VERSION : 0.1
   VAR_INPUT
      CMD : Bool;   // Команда запуска
      Res_1 : DInt;   // Наработка устройства 1
      Res_2 : DInt;   // Наработка устройства 2
      Alm_1 : Bool;   // Авария устройства 1
      Alm_2 : Bool;   // Авария устройства 2
   END_VAR
   VAR_IN_OUT
      Res_SP : DInt;   // Переключение по наработке
      CMD_1 : Bool;   // Команда на устройство 1
      CMD_2 : Bool;   // Команда на устройство 2
   END_VAR
   VAR_TEMP
      N : Bool;   // Выбор устройства
      Now : DInt;   // Текущая разница наработок
   END_VAR
BEGIN

REGION Network 1: Подсчёт разницы наработки
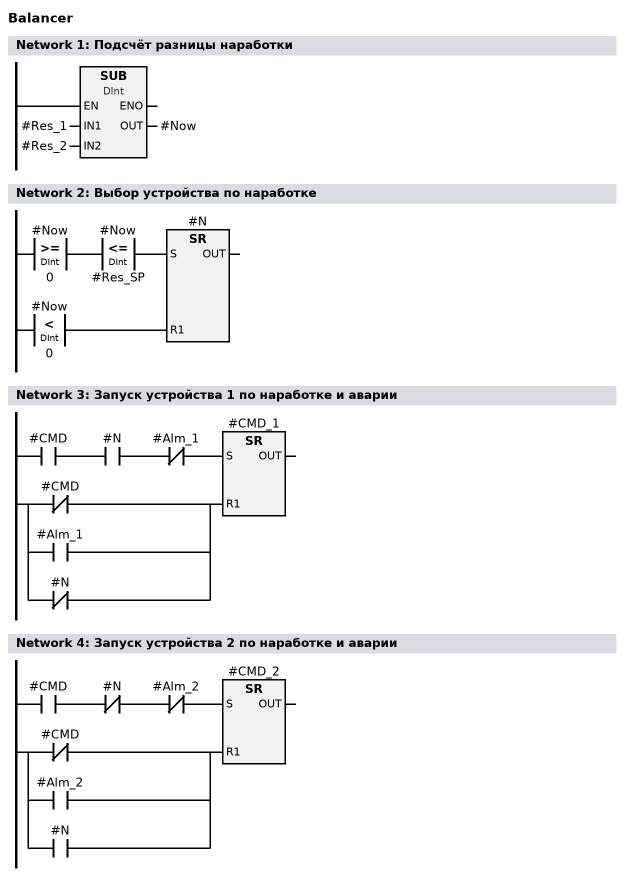
   RUNG wire#powerrail
      { S7_Templates := "SrcType := DInt"; S7_GenerateENO := "TRUE" } Sub(in1 := #Res_1, in2 := #Res_2, out => #Now)
   END_RUNG
   // the same network as SCL:
   #Now := #Res_1 - #Res_2;
END_REGION

REGION Network 2: Выбор устройства по наработке
   RUNG wire#powerrail
      { S7_Templates := "SrcType := DInt" } GE_Contact(in1 := #Now, in2 := 0)
      { S7_Templates := "SrcType := DInt" } LE_Contact(in1 := #Now, in2 := #Res_SP)
      S_SR(operand := #N, r1 := wire#w1)
   END_RUNG
   RUNG wire#powerrail
      { S7_Templates := "SrcType := DInt" } LT_Contact(in1 := #Now, in2 := 0)
   END_RUNG wire#w1
   // the same network as SCL:
   IF (#Now >= 0) AND (#Now <= #Res_SP) THEN
       #N := TRUE;   // SR flip-flop
   END_IF;
   IF #Now < 0 THEN #N := FALSE; END_IF;
END_REGION

REGION Network 3: Запуск устройства 1 по наработке и аварии
   RUNG wire#powerrail
      Contact( #CMD )
      Contact( #N )
      I_Contact( #Alm_1 )
      S_SR(operand := #CMD_1, r1 := wire#w1)
   END_RUNG
   RUNG wire#powerrail
      I_Contact( #CMD )
   END_RUNG wire#w1
   RUNG wire#powerrail
      Contact( #Alm_1 )
   END_RUNG wire#w1
   RUNG wire#powerrail
      I_Contact( #N )
   END_RUNG wire#w1
   // the same network as SCL:
   IF #CMD AND #N AND NOT #Alm_1 THEN
       #CMD_1 := TRUE;   // SR flip-flop
   END_IF;
   IF NOT #CMD OR #Alm_1 OR NOT #N THEN #CMD_1 := FALSE; END_IF;
END_REGION

REGION Network 4: Запуск устройства 2 по наработке и аварии
   RUNG wire#powerrail
      Contact( #CMD )
      I_Contact( #N )
      I_Contact( #Alm_2 )
      S_SR(operand := #CMD_2, r1 := wire#w1)
   END_RUNG
   RUNG wire#powerrail
      I_Contact( #CMD )
   END_RUNG wire#w1
   RUNG wire#powerrail
      Contact( #Alm_2 )
   END_RUNG wire#w1
   RUNG wire#powerrail
      Contact( #N )
   END_RUNG wire#w1
   // the same network as SCL:
   IF #CMD AND NOT #N AND NOT #Alm_2 THEN
       #CMD_2 := TRUE;   // SR flip-flop
   END_IF;
   IF NOT #CMD OR #Alm_2 OR #N THEN #CMD_2 := FALSE; END_IF;
END_REGION
END_FUNCTION

FUNCTION "INV" : Void   // FC111, LAD
{ S7_Optimized_Access := 'TRUE' }
VERSION : 0.1
   VAR_INPUT
      S : Bool;   // Сигнал
      I : Bool;   // Инверсия
   END_VAR
   VAR_IN_OUT
      R : Bool;   // Результат
   END_VAR
BEGIN

REGION Network 1: Инверсия сигнала
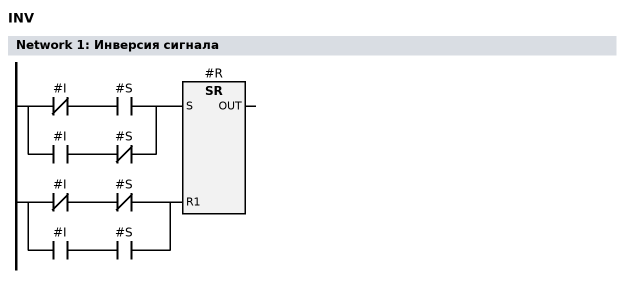
   RUNG wire#powerrail
      I_Contact( #I )
      Contact( #S )
      wire#w1
      S_SR(operand := #R, r1 := wire#w2)
   END_RUNG
   RUNG wire#powerrail
      Contact( #I )
      I_Contact( #S )
   END_RUNG wire#w1
   RUNG wire#powerrail
      I_Contact( #I )
      I_Contact( #S )
   END_RUNG wire#w2
   RUNG wire#powerrail
      Contact( #I )
      Contact( #S )
   END_RUNG wire#w2
   // the same network as SCL:
   IF (NOT #I AND #S) OR (#I AND NOT #S) THEN
       #R := TRUE;   // SR flip-flop
   END_IF;
   IF (NOT #I AND NOT #S) OR (#I AND #S) THEN #R := FALSE; END_IF;
END_REGION
END_FUNCTION

FUNCTION "Mode" : Void   // FC150, LAD
{ S7_Optimized_Access := 'FALSE' }
VERSION : 0.1
   VAR_INPUT
      CMD : Struct   // Основные команды
         Hand : Bool;   // 0 - авто, 1 - ручной / 0 - Авто, 1 - Ручной
         Start_A : Bool;   // Автозапуск / Запуск в авторежиме
         Start_M : Bool;   // Ручной - вперёд / Запуск в ручном режиме
         Force : Bool;   // Принудительный
         Lock : Bool;   // Блокировать / Блокировка
         Local : Bool;   // Локальный
         Service : Bool;   // Сервис
         Safety : Bool;   // Безопасность
         Alarm : Bool;   // Есть авария / Авария
         Reset : Bool;   // Сброс аварий
         Sim : Bool;   // Режим симуляции
      END_STRUCT;
      All_Block : Bool;   // Аварийная блокировка
   END_VAR
   VAR_OUTPUT
      Mode : Int;   // Режим работы
   END_VAR
BEGIN

REGION Network 1: Автоматический режим
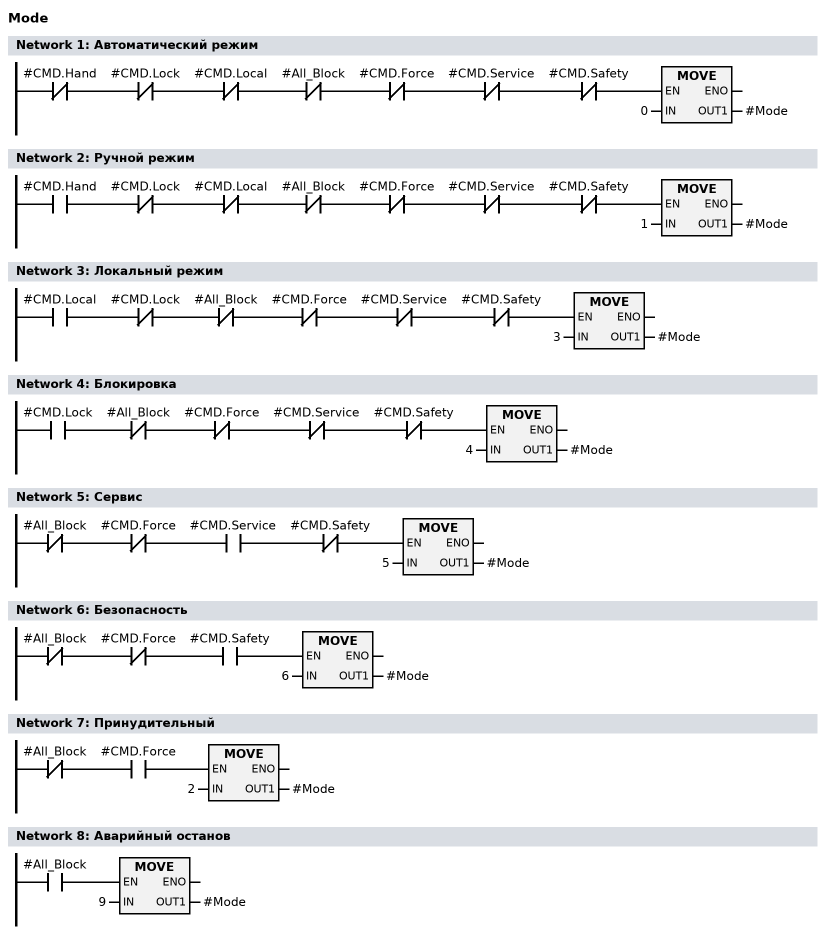
   RUNG wire#powerrail
      I_Contact( #CMD.Hand )
      I_Contact( #CMD.Lock )
      I_Contact( #CMD.Local )
      I_Contact( #All_Block )
      I_Contact( #CMD.Force )
      I_Contact( #CMD.Service )
      I_Contact( #CMD.Safety )
      { S7_GenerateENO := "TRUE" } Move(in := 0, out1 => #Mode)
   END_RUNG
   // the same network as SCL:
   IF NOT #CMD.Hand AND NOT #CMD.Lock AND NOT #CMD.Local AND NOT #All_Block AND NOT #CMD.Force AND NOT #CMD.Service AND NOT #CMD.Safety THEN
       #Mode := 0;
   END_IF;
END_REGION

REGION Network 2: Ручной режим
   RUNG wire#powerrail
      Contact( #CMD.Hand )
      I_Contact( #CMD.Lock )
      I_Contact( #CMD.Local )
      I_Contact( #All_Block )
      I_Contact( #CMD.Force )
      I_Contact( #CMD.Service )
      I_Contact( #CMD.Safety )
      { S7_GenerateENO := "TRUE" } Move(in := 1, out1 => #Mode)
   END_RUNG
   // the same network as SCL:
   IF #CMD.Hand AND NOT #CMD.Lock AND NOT #CMD.Local AND NOT #All_Block AND NOT #CMD.Force AND NOT #CMD.Service AND NOT #CMD.Safety THEN
       #Mode := 1;
   END_IF;
END_REGION

REGION Network 3: Локальный режим
   RUNG wire#powerrail
      Contact( #CMD.Local )
      I_Contact( #CMD.Lock )
      I_Contact( #All_Block )
      I_Contact( #CMD.Force )
      I_Contact( #CMD.Service )
      I_Contact( #CMD.Safety )
      { S7_GenerateENO := "TRUE" } Move(in := 3, out1 => #Mode)
   END_RUNG
   // the same network as SCL:
   IF #CMD.Local AND NOT #CMD.Lock AND NOT #All_Block AND NOT #CMD.Force AND NOT #CMD.Service AND NOT #CMD.Safety THEN
       #Mode := 3;
   END_IF;
END_REGION

REGION Network 4: Блокировка
   RUNG wire#powerrail
      Contact( #CMD.Lock )
      I_Contact( #All_Block )
      I_Contact( #CMD.Force )
      I_Contact( #CMD.Service )
      I_Contact( #CMD.Safety )
      { S7_GenerateENO := "TRUE" } Move(in := 4, out1 => #Mode)
   END_RUNG
   // the same network as SCL:
   IF #CMD.Lock AND NOT #All_Block AND NOT #CMD.Force AND NOT #CMD.Service AND NOT #CMD.Safety THEN
       #Mode := 4;
   END_IF;
END_REGION

REGION Network 5: Сервис
   RUNG wire#powerrail
      I_Contact( #All_Block )
      I_Contact( #CMD.Force )
      Contact( #CMD.Service )
      I_Contact( #CMD.Safety )
      { S7_GenerateENO := "TRUE" } Move(in := 5, out1 => #Mode)
   END_RUNG
   // the same network as SCL:
   IF NOT #All_Block AND NOT #CMD.Force AND #CMD.Service AND NOT #CMD.Safety THEN #Mode := 5; END_IF;
END_REGION

REGION Network 6: Безопасность
   RUNG wire#powerrail
      I_Contact( #All_Block )
      I_Contact( #CMD.Force )
      Contact( #CMD.Safety )
      { S7_GenerateENO := "TRUE" } Move(in := 6, out1 => #Mode)
   END_RUNG
   // the same network as SCL:
   IF NOT #All_Block AND NOT #CMD.Force AND #CMD.Safety THEN #Mode := 6; END_IF;
END_REGION

REGION Network 7: Принудительный
   RUNG wire#powerrail
      I_Contact( #All_Block )
      Contact( #CMD.Force )
      { S7_GenerateENO := "TRUE" } Move(in := 2, out1 => #Mode)
   END_RUNG
   // the same network as SCL:
   IF NOT #All_Block AND #CMD.Force THEN #Mode := 2; END_IF;
END_REGION

REGION Network 8: Аварийный останов
   RUNG wire#powerrail
      Contact( #All_Block )
      { S7_GenerateENO := "TRUE" } Move(in := 9, out1 => #Mode)
   END_RUNG
   // the same network as SCL:
   IF #All_Block THEN #Mode := 9; END_IF;
END_REGION
END_FUNCTION

// ===== PLC "PLC_PolyMix_002"  CPU 1214C DC/DC/DC =====
// protected blocks, not shown: "AI_ex", "AIx", "AO_ex", "DRV_M_D", "FlowMeter", "Logick", "Motors", "PLF_FC", "Time_m", "Time_r", "Time_s"

VAR_GLOBAL   // PLC tag table "Default tag table"
   "Mix_1_Clock" AT %M10.0 : Bool;
   "Mix_2_Clock" AT %M10.1 : Bool;
   "Mix_3_Clock" AT %M10.2 : Bool;
   "Flow" AT %IW256 : Int;
   "Level" AT %IW258 : Int;
END_VAR

VAR_GLOBAL   // PLC tag table "Sys"
   "pulse_01s" AT %M2.0 : Bool;
   "pulse_05s" AT %M2.1 : Bool;
   "pulse_1s" AT %M2.2 : Bool;
   "All_block" AT %M3.0 : Bool;
   "Reset_All" AT %M3.1 : Bool;
   "Sim_All" AT %M3.2 : Bool;
   "Any_Hand" AT %M5.0 : Bool;
   "DI_Hand" AT %M5.1 : Bool;
   "DO_Hand" AT %M5.2 : Bool;
   "AI_Hand" AT %M5.3 : Bool;
   "AO_Hand" AT %M5.4 : Bool;
   "M_Hand" AT %M5.5 : Bool;
   "V_Hand" AT %M5.6 : Bool;
   "X_Hand" AT %M5.7 : Bool;
   "System_Byte" AT %MB1 : Byte;
   "FirstScan" AT %M1.0 : Bool;
   "DiagStatusUpdate" AT %M1.1 : Bool;
   "ON" AT %M1.2 : Bool;
   "OFF" AT %M1.3 : Bool;
   "Clock_Byte" AT %MB0 : Byte;
   "Clock_10Hz" AT %M0.0 : Bool;
   "Clock_5Hz" AT %M0.1 : Bool;
   "Clock_2.5Hz" AT %M0.2 : Bool;
   "Clock_2Hz" AT %M0.3 : Bool;
   "Clock_1.25Hz" AT %M0.4 : Bool;
   "Clock_1Hz" AT %M0.5 : Bool;
   "Clock_0.625Hz" AT %M0.6 : Bool;
   "Clock_0.5Hz" AT %M0.7 : Bool;
   "F_pulse_01s" AT %M2.3 : Bool;
   "F_pulse_05s" AT %M2.4 : Bool;
   "F_pulse_1s" AT %M2.5 : Bool;
   "FN_pulse_01s" AT %M2.6 : Bool;
   "Clock_5s" AT %M2.7 : Bool;
   "Any_Alm" AT %M6.0 : Bool;
   "AI_Alm" AT %M6.1 : Bool;
   "M_Alm" AT %M6.2 : Bool;
   "V_Alm" AT %M6.3 : Bool;
   "C_Alm" AT %M6.4 : Bool;
   "N_Alm" AT %M6.5 : Bool;
   "L_Alm" AT %M6.6 : Bool;
   "X_Alm" AT %M6.7 : Bool;
END_VAR

VAR_GLOBAL   // PLC tag table "IO Table"
   "DD_FB_Ready" AT %I0.6 : Bool;   // I 0.6 - Дозатор сухого вещества - готовность
   "Dos_FB_Run" AT %I0.7 : Bool;   // I 0.7 - Дозатор - работа
   "DD_LLS" AT %I1.0 : Bool;   // I 1.0 - Дозатор сухого вещества - низкий уровень
   "Vibro_FB_Ready" AT %I1.1 : Bool;   // I 1.1 - Вибратор - готовность
   "Transporter" AT %I1.2 : Bool;   // I 1.2 - Пневмотранспортёр - готовность
   "DL_FB_Ready" AT %I1.3 : Bool;   // I 1.3 - Дозатор жидкого вещества - готовность
   "Dry_Run" AT %I1.4 : Bool;   // I 1.4 - Датчик протока
   "AllBlock" AT %I1.5 : Bool;   // I 1.5 - Датчик перелива или Аварийная остановка
   "M1_FB_Ready" AT %I0.0 : Bool;   // I 0.0 - Мешалка 1 - готовность
   "M1_FB_Run" AT %I0.1 : Bool;   // I 0.1 - Мешалка 1 - работа
   "M2_FB_Ready" AT %I0.2 : Bool;   // I 0.2 - Мешалка 2 - готовность
   "M2_FB_Run" AT %I0.3 : Bool;   // I 0.3 - Мешалка 2 - работа
   "M3_FB_Ready" AT %I0.4 : Bool;   // I 0.4 - Мешалка 3 - готовность
   "M3_FB_Run" AT %I0.5 : Bool;   // I 0.5 - Мешалка 3 - работа
   "M1_CMD" AT %Q0.0 : Bool;   // Q 0.0 - Мешалка 1 - запуск
   "M2_CMD" AT %Q0.1 : Bool;   // Q 0.1 - Мешалка 2 - запуск
   "M3_CMD" AT %Q0.2 : Bool;   // Q 0.2 - Мешалка 3 - запуск
   "DD_CMD" AT %Q0.3 : Bool;   // Q 0.3 - Дозатор сухого вещества - запуск
   "Vibro_CMD" AT %Q0.4 : Bool;   // Q 0.4 - Вибратор - запуск
   "DL_CMD" AT %Q0.5 : Bool;   // Q 0.5 - Дозатор жидкого вещества - запуск
   "KC1_CMD" AT %Q0.6 : Bool;   // Q 0.6 - Соленоидный клапан КС1
   "LED_Dry_Run" AT %Q0.7 : Bool;   // Q 0.7 - LED - сухой ход
   "LED_Alarm" AT %Q1.0 : Bool;   // Q 1.0 - LED - общая авария
   "LED_Empty" AT %Q1.1 : Bool;   // Q 1.1 - LED - бункер пуст
END_VAR

DATA_BLOCK "Any_DB"   // DB3
{ S7_Optimized_Access := 'FALSE' }
VERSION : 0.1
   VAR
      Level_M : Int;
      Level_S : Int;
      Flow_M : Int;
      Flow_S : Int;
      DD_View : Bool;
      Level_View : Bool;
   END_VAR
BEGIN
END_DATA_BLOCK

DATA_BLOCK "CONFIG"   // DB10
{ S7_Optimized_Access := 'FALSE' }
VERSION : 0.1
   VAR
      Config : Struct
         Use_DD : Bool;   // Использовать сухой дозатор
         Use_DL : Bool := true;   // Использовать жидкий дозатор
         Use_Mix_1 : Bool := true;   // Использовать мешалку 1
         Use_Mix_2 : Bool := true;   // Использовать мешалку 2
         Use_Mix_3 : Bool := true;   // Использовать мешалку 3
      END_STRUCT;
   END_VAR
BEGIN
END_DATA_BLOCK

DATA_BLOCK "Comm_DB"   // DB11
{ S7_Optimized_Access := 'FALSE' }
VERSION : 0.1
   VAR
      DD_Status : Int;
      DD_Mode : Int;
      DD_Alarm : Word;
      DL_Status : Int;
      DL_Mode : Int;
      DL_Alarm : Word;
      Mix_1_Status : Int;
      Mix_1_Mode : Int;
      Mix_1_Alarm : Word;
      Mix_2_Status : Int;
      Mix_2_Mode : Int;
      Mix_2_Alarm : Word;
      Mix_3_Status : Int;
      Mix_3_Mode : Int;
      Mix_3_Alarm : Word;
      KC1_Status : Int;
      Flowmeter : Real;
      Flow_Alarm : Word;
      Level : Real;
      Level_Alarm : Word;
      SP : Real;
      Start : Bool;
      Hand : Bool;
      Warning : Bool;
      Config : Struct
         Use_DD : Bool;   // Использовать сухой дозатор
         Use_DL : Bool;   // Использовать жидкий дозатор
         Use_Mix_1 : Bool;   // Использовать мешалку 1
         Use_Mix_2 : Bool;   // Использовать мешалку 2
         Use_Mix_3 : Bool;   // Использовать мешалку 3
      END_STRUCT;
      Alarm : Word;
   END_VAR
BEGIN
END_DATA_BLOCK

// folder: Modules

DATA_BLOCK "DIx_DB"   // DB200
{ S7_Optimized_Access := 'FALSE' }
VERSION : 0.1
// stored: InstanceOfName DIx
"DIx"
BEGIN
END_DATA_BLOCK

DATA_BLOCK "DOx_DB"   // DB201
{ S7_Optimized_Access := 'FALSE' }
VERSION : 0.1
// stored: InstanceOfName DOx
"DOx"
BEGIN
END_DATA_BLOCK

DATA_BLOCK "Micro_DB"   // DB207
{ S7_Optimized_Access := 'FALSE' }
VERSION : 0.1
// stored: InstanceOfName Micro
"Micro"
BEGIN
END_DATA_BLOCK

// folder: System blocks/Program resources

DATA_BLOCK "T_Reset"   // DB7
{ S7_Optimized_Access := 'TRUE' }
AUTHOR : Simatic
FAMILY : IEC
NAME : IEC_TMR
VERSION : 1.0
// stored: InstanceOfName IEC_TIMER
"IEC_TIMER"
BEGIN
END_DATA_BLOCK

DATA_BLOCK "clock_5s_ON"   // DB507
{ S7_Optimized_Access := 'TRUE' }
AUTHOR : Simatic
FAMILY : IEC
NAME : IEC_TMR
VERSION : 1.0
// stored: InstanceOfName IEC_TIMER
"IEC_TIMER"
BEGIN
END_DATA_BLOCK

DATA_BLOCK "clock_5s_OFF"   // DB508
{ S7_Optimized_Access := 'TRUE' }
AUTHOR : Simatic
FAMILY : IEC
NAME : IEC_TMR
VERSION : 1.0
// stored: InstanceOfName IEC_TIMER
"IEC_TIMER"
BEGIN
END_DATA_BLOCK

// folder: (top level)

FUNCTION "Comm_FC" : Void   // FC1, LAD
{ S7_Optimized_Access := 'TRUE' }
VERSION : 0.1
BEGIN

REGION Network 1: Сухой дозатор
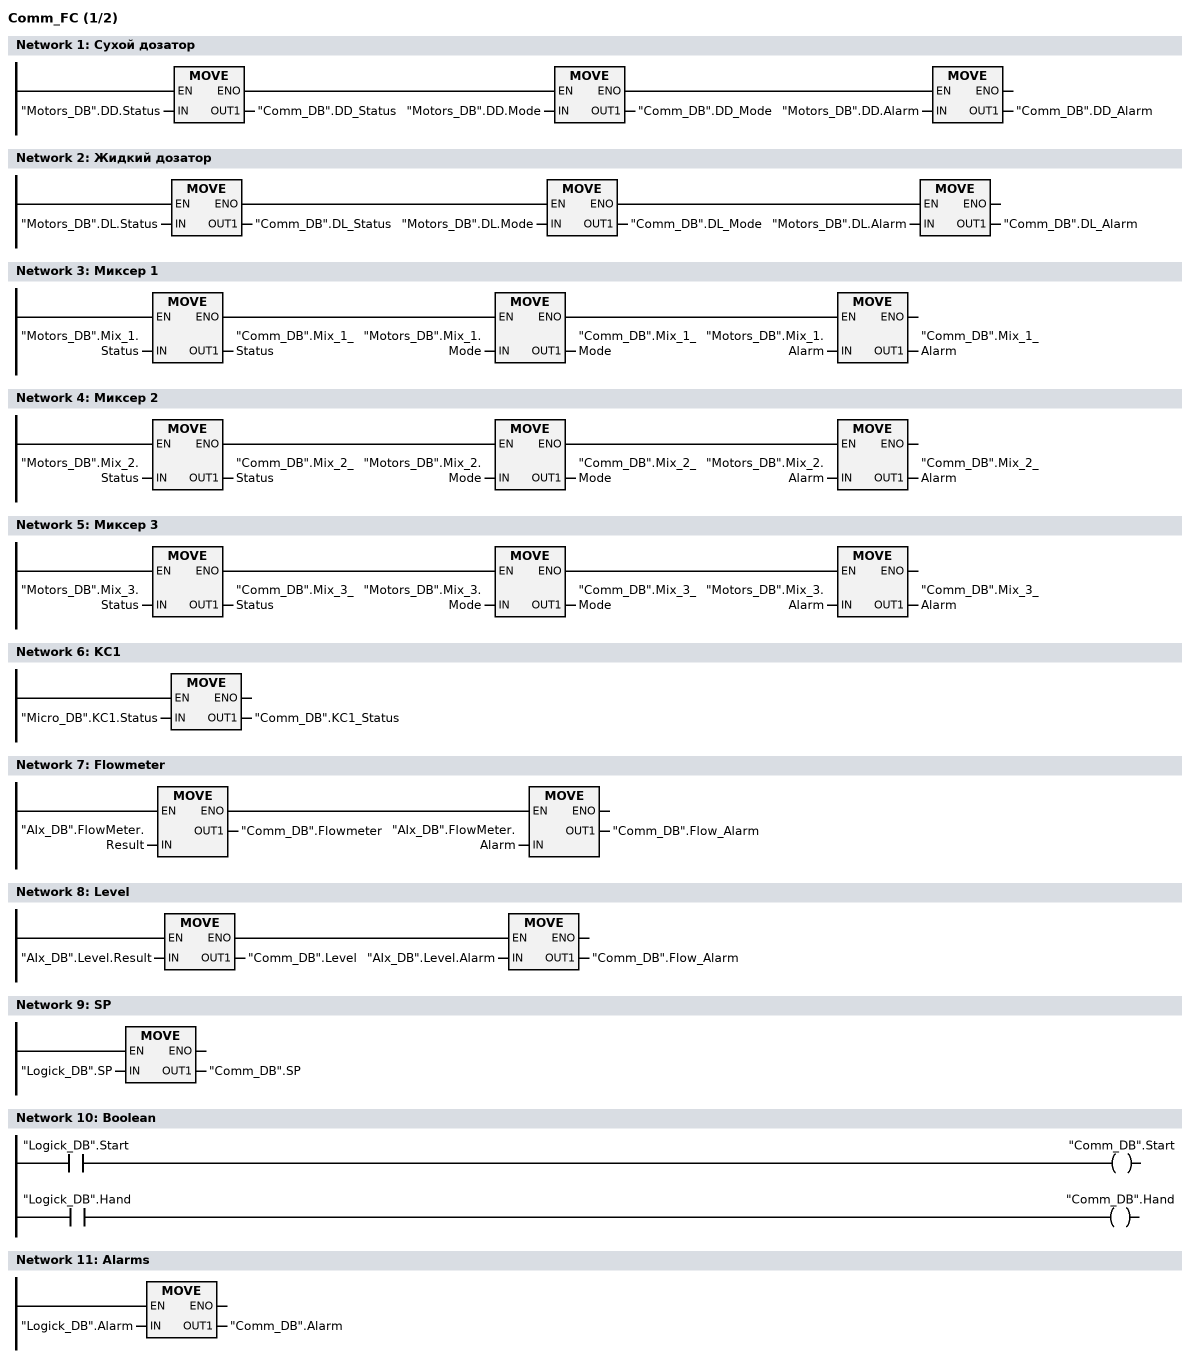
   RUNG wire#powerrail
      Move(in := "Motors_DB".DD.Status, out1 => "Comm_DB".DD_Status)
      Move(in := "Motors_DB".DD.Mode, out1 => "Comm_DB".DD_Mode)
      Move(in := "Motors_DB".DD.Alarm, out1 => "Comm_DB".DD_Alarm)
   END_RUNG
   // the same network as SCL:
   "Comm_DB".DD_Status := "Motors_DB".DD.Status;
   "Comm_DB".DD_Mode := "Motors_DB".DD.Mode;
   "Comm_DB".DD_Alarm := "Motors_DB".DD.Alarm;
END_REGION

REGION Network 2: Жидкий дозатор
   RUNG wire#powerrail
      Move(in := "Motors_DB".DL.Status, out1 => "Comm_DB".DL_Status)
      Move(in := "Motors_DB".DL.Mode, out1 => "Comm_DB".DL_Mode)
      Move(in := "Motors_DB".DL.Alarm, out1 => "Comm_DB".DL_Alarm)
   END_RUNG
   // the same network as SCL:
   "Comm_DB".DL_Status := "Motors_DB".DL.Status;
   "Comm_DB".DL_Mode := "Motors_DB".DL.Mode;
   "Comm_DB".DL_Alarm := "Motors_DB".DL.Alarm;
END_REGION

REGION Network 3: Миксер 1
   RUNG wire#powerrail
      Move(in := "Motors_DB".Mix_1.Status, out1 => "Comm_DB".Mix_1_Status)
      Move(in := "Motors_DB".Mix_1.Mode, out1 => "Comm_DB".Mix_1_Mode)
      Move(in := "Motors_DB".Mix_1.Alarm, out1 => "Comm_DB".Mix_1_Alarm)
   END_RUNG
   // the same network as SCL:
   "Comm_DB".Mix_1_Status := "Motors_DB".Mix_1.Status;
   "Comm_DB".Mix_1_Mode := "Motors_DB".Mix_1.Mode;
   "Comm_DB".Mix_1_Alarm := "Motors_DB".Mix_1.Alarm;
END_REGION

REGION Network 4: Миксер 2
   RUNG wire#powerrail
      Move(in := "Motors_DB".Mix_2.Status, out1 => "Comm_DB".Mix_2_Status)
      Move(in := "Motors_DB".Mix_2.Mode, out1 => "Comm_DB".Mix_2_Mode)
      Move(in := "Motors_DB".Mix_2.Alarm, out1 => "Comm_DB".Mix_2_Alarm)
   END_RUNG
   // the same network as SCL:
   "Comm_DB".Mix_2_Status := "Motors_DB".Mix_2.Status;
   "Comm_DB".Mix_2_Mode := "Motors_DB".Mix_2.Mode;
   "Comm_DB".Mix_2_Alarm := "Motors_DB".Mix_2.Alarm;
END_REGION

REGION Network 5: Миксер 3
   RUNG wire#powerrail
      Move(in := "Motors_DB".Mix_3.Status, out1 => "Comm_DB".Mix_3_Status)
      Move(in := "Motors_DB".Mix_3.Mode, out1 => "Comm_DB".Mix_3_Mode)
      Move(in := "Motors_DB".Mix_3.Alarm, out1 => "Comm_DB".Mix_3_Alarm)
   END_RUNG
   // the same network as SCL:
   "Comm_DB".Mix_3_Status := "Motors_DB".Mix_3.Status;
   "Comm_DB".Mix_3_Mode := "Motors_DB".Mix_3.Mode;
   "Comm_DB".Mix_3_Alarm := "Motors_DB".Mix_3.Alarm;
END_REGION

REGION Network 6: KC1
   RUNG wire#powerrail
      Move(in := "Micro_DB".KC1.Status, out1 => "Comm_DB".KC1_Status)
   END_RUNG
   // the same network as SCL:
   "Comm_DB".KC1_Status := "Micro_DB".KC1.Status;
END_REGION

REGION Network 7: Flowmeter
   RUNG wire#powerrail
      Move(in := "AIx_DB".FlowMeter.Result, out1 => "Comm_DB".Flowmeter)
      Move(in := "AIx_DB".FlowMeter.Alarm, out1 => "Comm_DB".Flow_Alarm)
   END_RUNG
   // the same network as SCL:
   "Comm_DB".Flowmeter := "AIx_DB".FlowMeter.Result;
   "Comm_DB".Flow_Alarm := "AIx_DB".FlowMeter.Alarm;
END_REGION

REGION Network 8: Level
   RUNG wire#powerrail
      Move(in := "AIx_DB".Level.Result, out1 => "Comm_DB".Level)
      Move(in := "AIx_DB".Level.Alarm, out1 => "Comm_DB".Flow_Alarm)
   END_RUNG
   // the same network as SCL:
   "Comm_DB".Level := "AIx_DB".Level.Result;
   "Comm_DB".Flow_Alarm := "AIx_DB".Level.Alarm;
END_REGION

REGION Network 9: SP
   RUNG wire#powerrail
      Move(in := "Logick_DB".SP, out1 => "Comm_DB".SP)
   END_RUNG
   // the same network as SCL:
   "Comm_DB".SP := "Logick_DB".SP;
END_REGION

REGION Network 10: Boolean
   RUNG wire#powerrail
      Contact( "Logick_DB".Start )
      Coil( "Comm_DB".Start )
   END_RUNG
   RUNG wire#powerrail
      Contact( "Logick_DB".Hand )
      Coil( "Comm_DB".Hand )
   END_RUNG
   // the same network as SCL:
   "Comm_DB".Start := "Logick_DB".Start;
   "Comm_DB".Hand := "Logick_DB".Hand;
END_REGION

REGION Network 11: Alarms
   RUNG wire#powerrail
      Move(in := "Logick_DB".Alarm, out1 => "Comm_DB".Alarm)
   END_RUNG
   // the same network as SCL:
   "Comm_DB".Alarm := "Logick_DB".Alarm;
END_REGION

REGION Network 12: Config
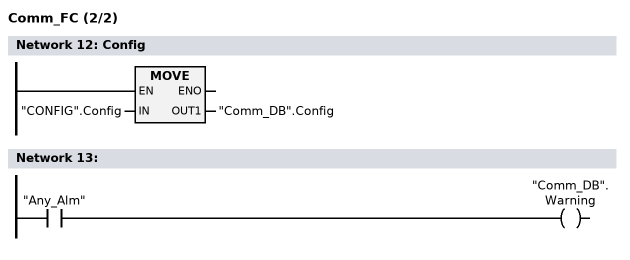
   RUNG wire#powerrail
      Move(in := "CONFIG".Config, out1 => "Comm_DB".Config)
   END_RUNG
   // the same network as SCL:
   "Comm_DB".Config := "CONFIG".Config;
END_REGION

REGION Network 13
   RUNG wire#powerrail
      Contact( "Any_Alm" )
      Coil( "Comm_DB".Warning )
   END_RUNG
   // the same network as SCL:
   "Comm_DB".Warning := "Any_Alm";
END_REGION
END_FUNCTION

ORGANIZATION_BLOCK "Main"   // OB1, LAD, ProgramCycle
TITLE = "Main Program Sweep (Cycle)"
{ S7_Optimized_Access := 'TRUE' }
VERSION : 0.1
   VAR_INPUT
      Initial_Call : Bool;   // Initial call of this OB
      Remanence : Bool;   // =True, if remanent data are available
   END_VAR
   VAR_TEMP   // added for the SCL form of the ladder/FBD networks
      _w1 : Bool;
   END_VAR
BEGIN

REGION Network 1
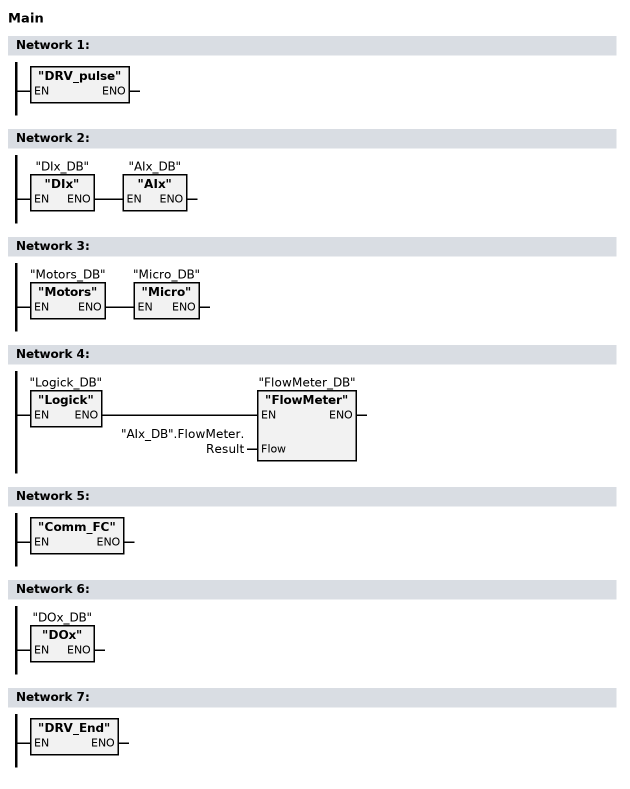
   RUNG wire#powerrail
      "DRV_pulse"()
   END_RUNG
   // the same network as SCL:
   "DRV_pulse"();
END_REGION

REGION Network 2
   RUNG wire#powerrail
      "DIx_DB"()
      "AIx_DB"()
   END_RUNG
   // the same network as SCL:
   "DIx_DB"(ENO => #_w1);   // "DIx"
   IF #_w1 THEN
       "AIx_DB"();   // "AIx"
   END_IF;
END_REGION

REGION Network 3
   RUNG wire#powerrail
      "Motors_DB"()
      "Micro_DB"()
   END_RUNG
   // the same network as SCL:
   "Motors_DB"(ENO => #_w1);   // "Motors"
   IF #_w1 THEN
       "Micro_DB"();   // "Micro"
   END_IF;
END_REGION

REGION Network 4
   RUNG wire#powerrail
      "Logick_DB"()
      "FlowMeter_DB"(Flow := "AIx_DB".FlowMeter.Result)
   END_RUNG
   // the same network as SCL:
   "Logick_DB"(ENO => #_w1);   // "Logick"
   IF #_w1 THEN
       "FlowMeter_DB"(Flow := "AIx_DB".FlowMeter.Result);   // "FlowMeter"
   END_IF;
END_REGION

REGION Network 5
   RUNG wire#powerrail
      "Comm_FC"()
   END_RUNG
   // the same network as SCL:
   "Comm_FC"();
END_REGION

REGION Network 6
   RUNG wire#powerrail
      "DOx_DB"()
   END_RUNG
   // the same network as SCL:
   "DOx_DB"();   // "DOx"
END_REGION

REGION Network 7
   RUNG wire#powerrail
      "DRV_End"()
   END_RUNG
   // the same network as SCL:
   "DRV_End"();
END_REGION
END_ORGANIZATION_BLOCK

ORGANIZATION_BLOCK "Time error interrupt"   // OB80, LAD, TimeErrorInterrupt
{ S7_Optimized_Access := 'TRUE' }
VERSION : 0.1
   VAR_INPUT
      Fault_ID : Byte;   // Fault identifier
      Csg_OBnr : OB_Any;   // Number of OB causing the error
      Csg_Prio : UInt;   // Priority of OB causing the error
   END_VAR
BEGIN
END_ORGANIZATION_BLOCK

ORGANIZATION_BLOCK "Diagnostic error interrupt"   // OB82, LAD, DiagnosticErrorInterrupt
{ S7_Optimized_Access := 'TRUE' }
VERSION : 0.1
   VAR_INPUT
      IO_State : Word;   // IO state of the HW object
      LADDR : Hw_Any;   // Hardware identifier
      Channel : UInt;   // Channel number
      MultiError : Bool;   // =true if more than one error is present
   END_VAR
BEGIN
END_ORGANIZATION_BLOCK

ORGANIZATION_BLOCK "Startup"   // OB100, LAD, Startup
TITLE = "Complete Restart"
{ S7_Optimized_Access := 'TRUE' }
VERSION : 0.1
   VAR_INPUT
      LostRetentive : Bool;   // True if retentive data are lost
      LostRTC : Bool;   // True if date and time are lost
   END_VAR
BEGIN

REGION Network 1: Запуск автоматики
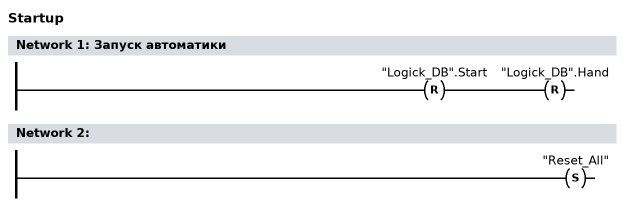
   RUNG wire#powerrail
      R_Coil( "Logick_DB".Start )
      R_Coil( "Logick_DB".Hand )
   END_RUNG
   // the same network as SCL:
   "Logick_DB".Start := FALSE;
   "Logick_DB".Hand := FALSE;
END_REGION

REGION Network 2
   RUNG wire#powerrail
      S_Coil( "Reset_All" )
   END_RUNG
   // the same network as SCL:
   "Reset_All" := TRUE;
END_REGION
END_ORGANIZATION_BLOCK

// folder: DRV_Low

FUNCTION_BLOCK "DI_ex"   // FB100, LAD
{ S7_Optimized_Access := 'FALSE' }
VERSION : 0.1
   VAR_INPUT
      Input : Bool;   // Входящий сигнал
      pulse : Bool;   // Частота фильтрации дребезка
   END_VAR
   VAR_OUTPUT
      Signal : Bool;   // Результирующий сигнал
   END_VAR
   VAR
      Hand : Bool;   // 0 - Авто, 1 - Ручной
      Start_M : Bool;   // Запуск в ручном режиме
      Data : Bool;   // Отфильтрованный сигнал
      Inverse : Bool;   // Инверсия входного сигнала
      Filter_On : Struct   // Фильтр наличия сигнала
         SP : Int;
         Now : Int;
         "Exit" : Bool;
         Start : Bool;
         Pause : Bool;
         Reset : Bool;
      END_STRUCT;
      Filter_Off : Struct   // Фильтр отсутствия сигнала
         SP : Int;
         Now : Int;
         "Exit" : Bool;
         Start : Bool;
         Pause : Bool;
         Reset : Bool;
      END_STRUCT;
      res_1 : Word;
   END_VAR
   VAR_TEMP   // added for the SCL form of the ladder/FBD networks
      _w1 : Bool;
   END_VAR
BEGIN

REGION Network 1: Устройство в ручном режиме
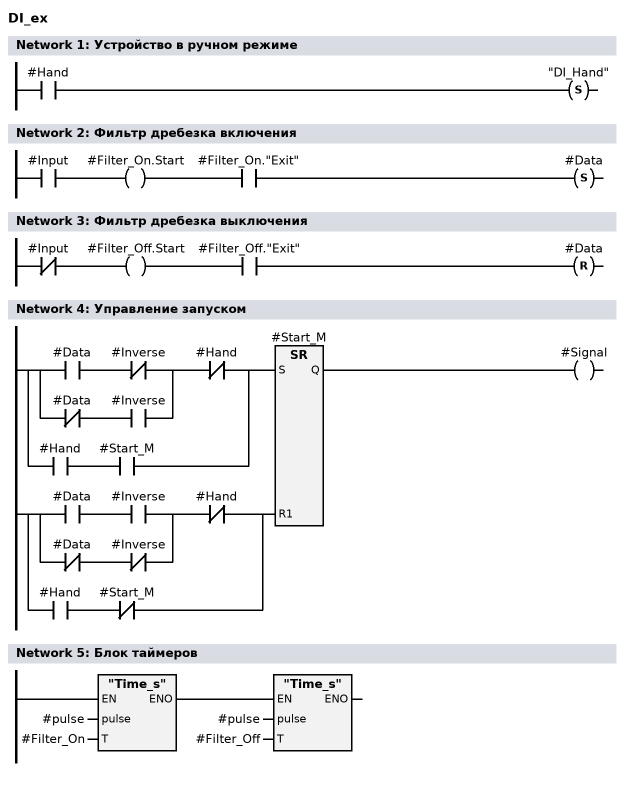
   RUNG wire#powerrail
      Contact( #Hand )
      S_Coil( "DI_Hand" )
   END_RUNG
   // the same network as SCL:
   IF #Hand THEN "DI_Hand" := TRUE; END_IF;
END_REGION

REGION Network 2: Фильтр дребезка включения
   RUNG wire#powerrail
      Contact( #Input )
      Coil( #Filter_On.Start )
      Contact( #Filter_On."Exit" )
      S_Coil( #Data )
   END_RUNG
   // the same network as SCL:
   #Filter_On.Start := #Input;
   IF #Input AND #Filter_On."Exit" THEN #Data := TRUE; END_IF;
END_REGION

REGION Network 3: Фильтр дребезка выключения
   RUNG wire#powerrail
      I_Contact( #Input )
      Coil( #Filter_Off.Start )
      Contact( #Filter_Off."Exit" )
      R_Coil( #Data )
   END_RUNG
   // the same network as SCL:
   #Filter_Off.Start := NOT #Input;
   IF NOT #Input AND #Filter_Off."Exit" THEN #Data := FALSE; END_IF;
END_REGION
